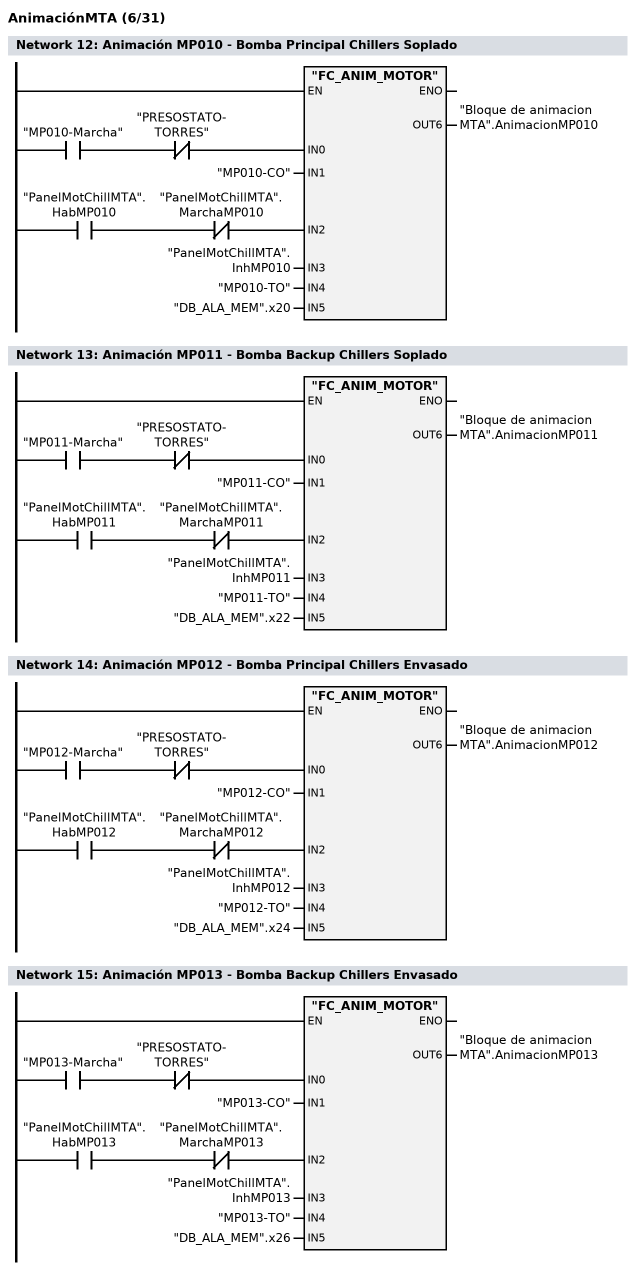
   RUNG wire#powerrail
      "FC_ANIM_MOTOR"(IN0 := wire#w1, IN2 := wire#w2, IN1 := "MP010-CO", IN3 := "PanelMotChillMTA".InhMP010, IN4 := "MP010-TO", IN5 := "DB_ALA_MEM".x20, OUT6 => "Bloque de animacion MTA".AnimacionMP010)
   END_RUNG
   RUNG wire#powerrail
      Contact( "MP010-Marcha" )
      I_Contact( "PRESOSTATO-TORRES" )
   END_RUNG wire#w1
   RUNG wire#powerrail
      Contact( "PanelMotChillMTA".HabMP010 )
      I_Contact( "PanelMotChillMTA".MarchaMP010 )
   END_RUNG wire#w2
   // the same network as SCL:
   "FC_ANIM_MOTOR"(IN0 := "MP010-Marcha" AND NOT "PRESOSTATO-TORRES",
                   IN1 := "MP010-CO",
                   IN2 := "PanelMotChillMTA".HabMP010 AND NOT "PanelMotChillMTA".MarchaMP010,
                   IN3 := "PanelMotChillMTA".InhMP010,
                   IN4 := "MP010-TO",
                   IN5 := "DB_ALA_MEM".x20,
                   OUT6 => "Bloque de animacion MTA".AnimacionMP010);
END_REGION

REGION Network 13: Animación MP011 - Bomba Backup Chillers Soplado
   RUNG wire#powerrail
      "FC_ANIM_MOTOR"(IN0 := wire#w1, IN2 := wire#w2, IN1 := "MP011-CO", IN3 := "PanelMotChillMTA".InhMP011, IN4 := "MP011-TO", IN5 := "DB_ALA_MEM".x22, OUT6 => "Bloque de animacion MTA".AnimacionMP011)
   END_RUNG
   RUNG wire#powerrail
      Contact( "MP011-Marcha" )
      I_Contact( "PRESOSTATO-TORRES" )
   END_RUNG wire#w1
   RUNG wire#powerrail
      Contact( "PanelMotChillMTA".HabMP011 )
      I_Contact( "PanelMotChillMTA".MarchaMP011 )
   END_RUNG wire#w2
   // the same network as SCL:
   "FC_ANIM_MOTOR"(IN0 := "MP011-Marcha" AND NOT "PRESOSTATO-TORRES",
                   IN1 := "MP011-CO",
                   IN2 := "PanelMotChillMTA".HabMP011 AND NOT "PanelMotChillMTA".MarchaMP011,
                   IN3 := "PanelMotChillMTA".InhMP011,
                   IN4 := "MP011-TO",
                   IN5 := "DB_ALA_MEM".x22,
                   OUT6 => "Bloque de animacion MTA".AnimacionMP011);
END_REGION

REGION Network 14: Animación MP012 - Bomba Principal Chillers Envasado
   RUNG wire#powerrail
      "FC_ANIM_MOTOR"(IN0 := wire#w1, IN2 := wire#w2, IN1 := "MP012-CO", IN3 := "PanelMotChillMTA".InhMP012, IN4 := "MP012-TO", IN5 := "DB_ALA_MEM".x24, OUT6 => "Bloque de animacion MTA".AnimacionMP012)
   END_RUNG
   RUNG wire#powerrail
      Contact( "MP012-Marcha" )
      I_Contact( "PRESOSTATO-TORRES" )
   END_RUNG wire#w1
   RUNG wire#powerrail
      Contact( "PanelMotChillMTA".HabMP012 )
      I_Contact( "PanelMotChillMTA".MarchaMP012 )
   END_RUNG wire#w2
   // the same network as SCL:
   "FC_ANIM_MOTOR"(IN0 := "MP012-Marcha" AND NOT "PRESOSTATO-TORRES",
                   IN1 := "MP012-CO",
                   IN2 := "PanelMotChillMTA".HabMP012 AND NOT "PanelMotChillMTA".MarchaMP012,
                   IN3 := "PanelMotChillMTA".InhMP012,
                   IN4 := "MP012-TO",
                   IN5 := "DB_ALA_MEM".x24,
                   OUT6 => "Bloque de animacion MTA".AnimacionMP012);
END_REGION

REGION Network 15: Animación MP013 - Bomba Backup Chillers Envasado
   RUNG wire#powerrail
      "FC_ANIM_MOTOR"(IN0 := wire#w1, IN2 := wire#w2, IN1 := "MP013-CO", IN3 := "PanelMotChillMTA".InhMP013, IN4 := "MP013-TO", IN5 := "DB_ALA_MEM".x26, OUT6 => "Bloque de animacion MTA".AnimacionMP013)
   END_RUNG
   RUNG wire#powerrail
      Contact( "MP013-Marcha" )
      I_Contact( "PRESOSTATO-TORRES" )
   END_RUNG wire#w1
   RUNG wire#powerrail
      Contact( "PanelMotChillMTA".HabMP013 )
      I_Contact( "PanelMotChillMTA".MarchaMP013 )
   END_RUNG wire#w2
   // the same network as SCL:
   "FC_ANIM_MOTOR"(IN0 := "MP013-Marcha" AND NOT "PRESOSTATO-TORRES",
                   IN1 := "MP013-CO",
                   IN2 := "PanelMotChillMTA".HabMP013 AND NOT "PanelMotChillMTA".MarchaMP013,
                   IN3 := "PanelMotChillMTA".InhMP013,
                   IN4 := "MP013-TO",
                   IN5 := "DB_ALA_MEM".x26,
                   OUT6 => "Bloque de animacion MTA".AnimacionMP013);
END_REGION

REGION Network 16: Animación MP018 - Bomba 1 Torres de enfriamiento
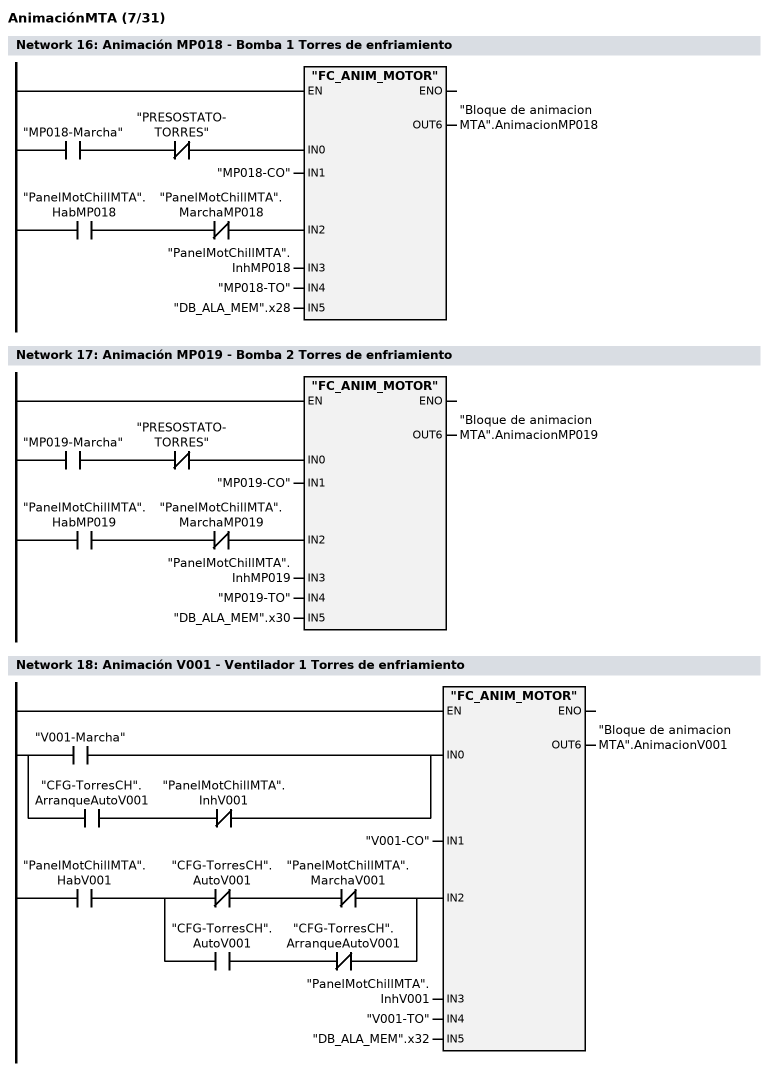
   RUNG wire#powerrail
      "FC_ANIM_MOTOR"(IN0 := wire#w1, IN2 := wire#w2, IN1 := "MP018-CO", IN3 := "PanelMotChillMTA".InhMP018, IN4 := "MP018-TO", IN5 := "DB_ALA_MEM".x28, OUT6 => "Bloque de animacion MTA".AnimacionMP018)
   END_RUNG
   RUNG wire#powerrail
      Contact( "MP018-Marcha" )
      I_Contact( "PRESOSTATO-TORRES" )
   END_RUNG wire#w1
   RUNG wire#powerrail
      Contact( "PanelMotChillMTA".HabMP018 )
      I_Contact( "PanelMotChillMTA".MarchaMP018 )
   END_RUNG wire#w2
   // the same network as SCL:
   "FC_ANIM_MOTOR"(IN0 := "MP018-Marcha" AND NOT "PRESOSTATO-TORRES",
                   IN1 := "MP018-CO",
                   IN2 := "PanelMotChillMTA".HabMP018 AND NOT "PanelMotChillMTA".MarchaMP018,
                   IN3 := "PanelMotChillMTA".InhMP018,
                   IN4 := "MP018-TO",
                   IN5 := "DB_ALA_MEM".x28,
                   OUT6 => "Bloque de animacion MTA".AnimacionMP018);
END_REGION

REGION Network 17: Animación MP019 - Bomba 2 Torres de enfriamiento
   RUNG wire#powerrail
      "FC_ANIM_MOTOR"(IN0 := wire#w1, IN2 := wire#w2, IN1 := "MP019-CO", IN3 := "PanelMotChillMTA".InhMP019, IN4 := "MP019-TO", IN5 := "DB_ALA_MEM".x30, OUT6 => "Bloque de animacion MTA".AnimacionMP019)
   END_RUNG
   RUNG wire#powerrail
      Contact( "MP019-Marcha" )
      I_Contact( "PRESOSTATO-TORRES" )
   END_RUNG wire#w1
   RUNG wire#powerrail
      Contact( "PanelMotChillMTA".HabMP019 )
      I_Contact( "PanelMotChillMTA".MarchaMP019 )
   END_RUNG wire#w2
   // the same network as SCL:
   "FC_ANIM_MOTOR"(IN0 := "MP019-Marcha" AND NOT "PRESOSTATO-TORRES",
                   IN1 := "MP019-CO",
                   IN2 := "PanelMotChillMTA".HabMP019 AND NOT "PanelMotChillMTA".MarchaMP019,
                   IN3 := "PanelMotChillMTA".InhMP019,
                   IN4 := "MP019-TO",
                   IN5 := "DB_ALA_MEM".x30,
                   OUT6 => "Bloque de animacion MTA".AnimacionMP019);
END_REGION

REGION Network 18: Animación V001 - Ventilador 1 Torres de enfriamiento
   RUNG wire#powerrail
      "FC_ANIM_MOTOR"(IN0 := wire#w1, IN2 := wire#w3, IN1 := "V001-CO", IN3 := "PanelMotChillMTA".InhV001, IN4 := "V001-TO", IN5 := "DB_ALA_MEM".x32, OUT6 => "Bloque de animacion MTA".AnimacionV001)
   END_RUNG
   RUNG wire#powerrail
      Contact( "V001-Marcha" )
   END_RUNG wire#w1
   RUNG wire#powerrail
      Contact( "CFG-TorresCH".ArranqueAutoV001 )
      I_Contact( "PanelMotChillMTA".InhV001 )
   END_RUNG wire#w1
   RUNG wire#powerrail
      Contact( "PanelMotChillMTA".HabV001 )
      wire#w2
      I_Contact( "CFG-TorresCH".AutoV001 )
      I_Contact( "PanelMotChillMTA".MarchaV001 )
   END_RUNG wire#w3
   RUNG wire#w2
      Contact( "CFG-TorresCH".AutoV001 )
      I_Contact( "CFG-TorresCH".ArranqueAutoV001 )
   END_RUNG wire#w3
   // the same network as SCL:
   "FC_ANIM_MOTOR"(IN0 := "V001-Marcha" OR ("CFG-TorresCH".ArranqueAutoV001 AND NOT "PanelMotChillMTA".InhV001),
                   IN1 := "V001-CO",
                   IN2 := "PanelMotChillMTA".HabV001 AND ((NOT "CFG-TorresCH".AutoV001 AND NOT "PanelMotChillMTA".MarchaV001) OR ("CFG-TorresCH".AutoV001 AND NOT "CFG-TorresCH".ArranqueAutoV001)),
                   IN3 := "PanelMotChillMTA".InhV001,
                   IN4 := "V001-TO",
                   IN5 := "DB_ALA_MEM".x32,
                   OUT6 => "Bloque de animacion MTA".AnimacionV001);
END_REGION

REGION Network 19: Animación V002 - Ventilador 2 Torres de enfriamiento
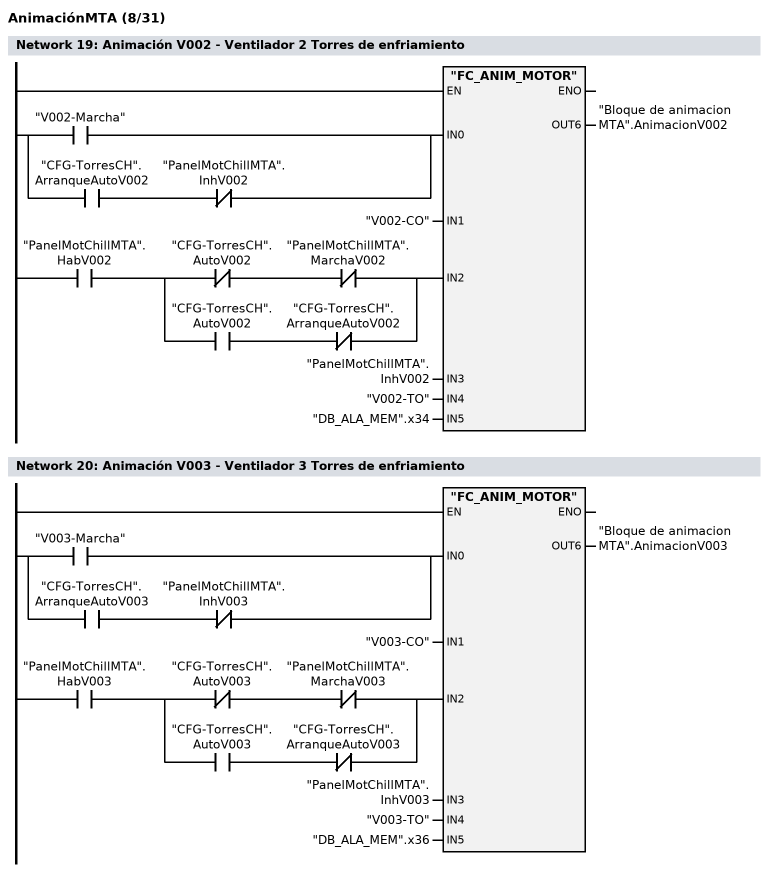
   RUNG wire#powerrail
      "FC_ANIM_MOTOR"(IN0 := wire#w1, IN2 := wire#w3, IN1 := "V002-CO", IN3 := "PanelMotChillMTA".InhV002, IN4 := "V002-TO", IN5 := "DB_ALA_MEM".x34, OUT6 => "Bloque de animacion MTA".AnimacionV002)
   END_RUNG
   RUNG wire#powerrail
      Contact( "V002-Marcha" )
   END_RUNG wire#w1
   RUNG wire#powerrail
      Contact( "CFG-TorresCH".ArranqueAutoV002 )
      I_Contact( "PanelMotChillMTA".InhV002 )
   END_RUNG wire#w1
   RUNG wire#powerrail
      Contact( "PanelMotChillMTA".HabV002 )
      wire#w2
      I_Contact( "CFG-TorresCH".AutoV002 )
      I_Contact( "PanelMotChillMTA".MarchaV002 )
   END_RUNG wire#w3
   RUNG wire#w2
      Contact( "CFG-TorresCH".AutoV002 )
      I_Contact( "CFG-TorresCH".ArranqueAutoV002 )
   END_RUNG wire#w3
   // the same network as SCL:
   "FC_ANIM_MOTOR"(IN0 := "V002-Marcha" OR ("CFG-TorresCH".ArranqueAutoV002 AND NOT "PanelMotChillMTA".InhV002),
                   IN1 := "V002-CO",
                   IN2 := "PanelMotChillMTA".HabV002 AND ((NOT "CFG-TorresCH".AutoV002 AND NOT "PanelMotChillMTA".MarchaV002) OR ("CFG-TorresCH".AutoV002 AND NOT "CFG-TorresCH".ArranqueAutoV002)),
                   IN3 := "PanelMotChillMTA".InhV002,
                   IN4 := "V002-TO",
                   IN5 := "DB_ALA_MEM".x34,
                   OUT6 => "Bloque de animacion MTA".AnimacionV002);
END_REGION

REGION Network 20: Animación V003 - Ventilador 3 Torres de enfriamiento
   RUNG wire#powerrail
      "FC_ANIM_MOTOR"(IN0 := wire#w1, IN2 := wire#w3, IN1 := "V003-CO", IN3 := "PanelMotChillMTA".InhV003, IN4 := "V003-TO", IN5 := "DB_ALA_MEM".x36, OUT6 => "Bloque de animacion MTA".AnimacionV003)
   END_RUNG
   RUNG wire#powerrail
      Contact( "V003-Marcha" )
   END_RUNG wire#w1
   RUNG wire#powerrail
      Contact( "CFG-TorresCH".ArranqueAutoV003 )
      I_Contact( "PanelMotChillMTA".InhV003 )
   END_RUNG wire#w1
   RUNG wire#powerrail
      Contact( "PanelMotChillMTA".HabV003 )
      wire#w2
      I_Contact( "CFG-TorresCH".AutoV003 )
      I_Contact( "PanelMotChillMTA".MarchaV003 )
   END_RUNG wire#w3
   RUNG wire#w2
      Contact( "CFG-TorresCH".AutoV003 )
      I_Contact( "CFG-TorresCH".ArranqueAutoV003 )
   END_RUNG wire#w3
   // the same network as SCL:
   "FC_ANIM_MOTOR"(IN0 := "V003-Marcha" OR ("CFG-TorresCH".ArranqueAutoV003 AND NOT "PanelMotChillMTA".InhV003),
                   IN1 := "V003-CO",
                   IN2 := "PanelMotChillMTA".HabV003 AND ((NOT "CFG-TorresCH".AutoV003 AND NOT "PanelMotChillMTA".MarchaV003) OR ("CFG-TorresCH".AutoV003 AND NOT "CFG-TorresCH".ArranqueAutoV003)),
                   IN3 := "PanelMotChillMTA".InhV003,
                   IN4 := "V003-TO",
                   IN5 := "DB_ALA_MEM".x36,
                   OUT6 => "Bloque de animacion MTA".AnimacionV003);
END_REGION

REGION Network 21: Animación MC060 - Compresor de Baja SULLAIR 2
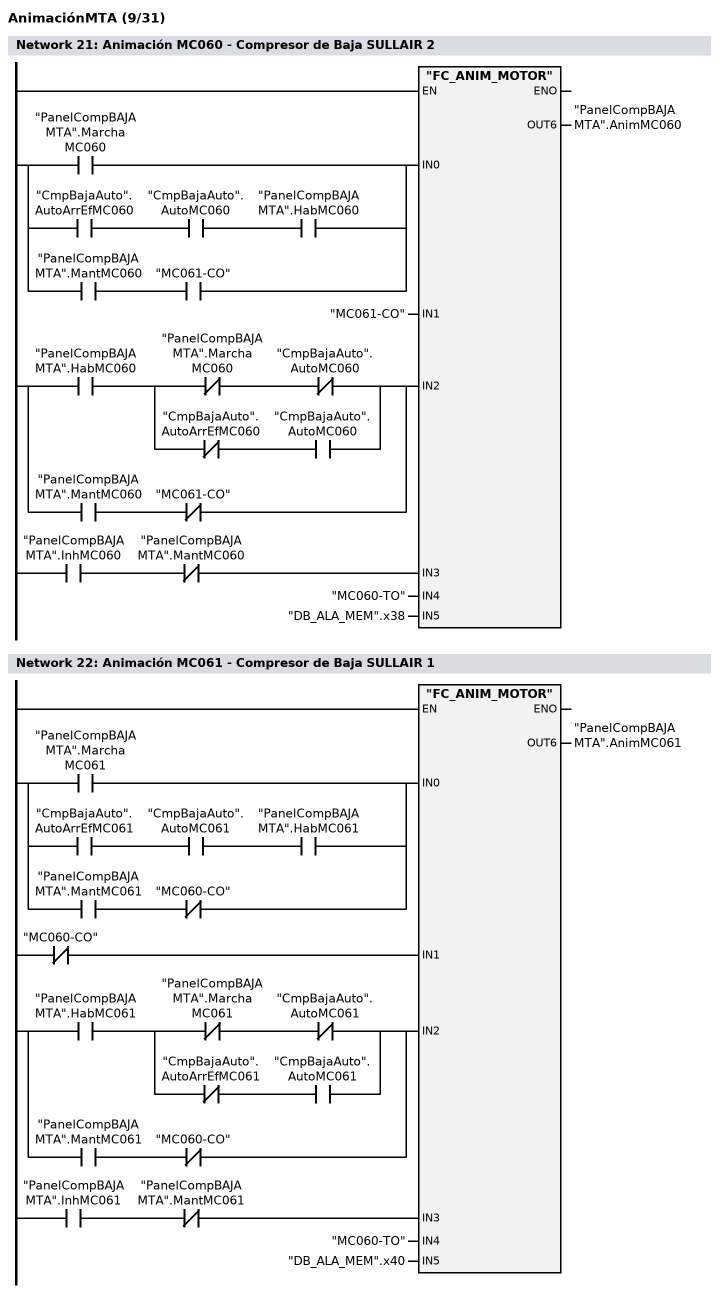
   RUNG wire#powerrail
      "FC_ANIM_MOTOR"(IN0 := wire#w1, IN2 := wire#w3, IN3 := wire#w4, IN1 := "MC061-CO", IN4 := "MC060-TO", IN5 := "DB_ALA_MEM".x38, OUT6 => "PanelCompBAJA MTA".AnimMC060)
   END_RUNG
   RUNG wire#powerrail
      Contact( "PanelCompBAJA MTA".MarchaMC060 )
   END_RUNG wire#w1
   RUNG wire#powerrail
      Contact( "CmpBajaAuto".AutoArrEfMC060 )
      Contact( "CmpBajaAuto".AutoMC060 )
      Contact( "PanelCompBAJA MTA".HabMC060 )
   END_RUNG wire#w1
   RUNG wire#powerrail
      Contact( "PanelCompBAJA MTA".MantMC060 )
      Contact( "MC061-CO" )
   END_RUNG wire#w1
   RUNG wire#powerrail
      Contact( "PanelCompBAJA MTA".HabMC060 )
      wire#w2
      I_Contact( "PanelCompBAJA MTA".MarchaMC060 )
      I_Contact( "CmpBajaAuto".AutoMC060 )
   END_RUNG wire#w3
   RUNG wire#w2
      I_Contact( "CmpBajaAuto".AutoArrEfMC060 )
      Contact( "CmpBajaAuto".AutoMC060 )
   END_RUNG wire#w3
   RUNG wire#powerrail
      Contact( "PanelCompBAJA MTA".MantMC060 )
      I_Contact( "MC061-CO" )
   END_RUNG wire#w3
   RUNG wire#powerrail
      Contact( "PanelCompBAJA MTA".InhMC060 )
      I_Contact( "PanelCompBAJA MTA".MantMC060 )
   END_RUNG wire#w4
   // the same network as SCL:
   "FC_ANIM_MOTOR"(IN0 := "PanelCompBAJA MTA".MarchaMC060 OR ("CmpBajaAuto".AutoArrEfMC060 AND "CmpBajaAuto".AutoMC060 AND "PanelCompBAJA MTA".HabMC060) OR ("PanelCompBAJA MTA".MantMC060 AND "MC061-CO"),
                   IN1 := "MC061-CO",
                   IN2 := ("PanelCompBAJA MTA".HabMC060 AND ((NOT "PanelCompBAJA MTA".MarchaMC060 AND NOT "CmpBajaAuto".AutoMC060) OR (NOT "CmpBajaAuto".AutoArrEfMC060 AND "CmpBajaAuto".AutoMC060))) OR ("PanelCompBAJA MTA".MantMC060 AND NOT "MC061-CO"),
                   IN3 := "PanelCompBAJA MTA".InhMC060 AND NOT "PanelCompBAJA MTA".MantMC060,
                   IN4 := "MC060-TO",
                   IN5 := "DB_ALA_MEM".x38,
                   OUT6 => "PanelCompBAJA MTA".AnimMC060);
END_REGION

REGION Network 22: Animación MC061 - Compresor de Baja SULLAIR 1
   RUNG wire#powerrail
      "FC_ANIM_MOTOR"(IN0 := wire#w1, IN1 := wire#w2, IN2 := wire#w4, IN3 := wire#w5, IN4 := "MC060-TO", IN5 := "DB_ALA_MEM".x40, OUT6 => "PanelCompBAJA MTA".AnimMC061)
   END_RUNG
   RUNG wire#powerrail
      Contact( "PanelCompBAJA MTA".MarchaMC061 )
   END_RUNG wire#w1
   RUNG wire#powerrail
      Contact( "CmpBajaAuto".AutoArrEfMC061 )
      Contact( "CmpBajaAuto".AutoMC061 )
      Contact( "PanelCompBAJA MTA".HabMC061 )
   END_RUNG wire#w1
   RUNG wire#powerrail
      Contact( "PanelCompBAJA MTA".MantMC061 )
      I_Contact( "MC060-CO" )
   END_RUNG wire#w1
   RUNG wire#powerrail
      I_Contact( "MC060-CO" )
   END_RUNG wire#w2
   RUNG wire#powerrail
      Contact( "PanelCompBAJA MTA".HabMC061 )
      wire#w3
      I_Contact( "PanelCompBAJA MTA".MarchaMC061 )
      I_Contact( "CmpBajaAuto".AutoMC061 )
   END_RUNG wire#w4
   RUNG wire#w3
      I_Contact( "CmpBajaAuto".AutoArrEfMC061 )
      Contact( "CmpBajaAuto".AutoMC061 )
   END_RUNG wire#w4
   RUNG wire#powerrail
      Contact( "PanelCompBAJA MTA".MantMC061 )
      I_Contact( "MC060-CO" )
   END_RUNG wire#w4
   RUNG wire#powerrail
      Contact( "PanelCompBAJA MTA".InhMC061 )
      I_Contact( "PanelCompBAJA MTA".MantMC061 )
   END_RUNG wire#w5
   // the same network as SCL:
   "FC_ANIM_MOTOR"(IN0 := "PanelCompBAJA MTA".MarchaMC061 OR ("CmpBajaAuto".AutoArrEfMC061 AND "CmpBajaAuto".AutoMC061 AND "PanelCompBAJA MTA".HabMC061) OR ("PanelCompBAJA MTA".MantMC061 AND NOT "MC060-CO"),
                   IN1 := NOT "MC060-CO",
                   IN2 := ("PanelCompBAJA MTA".HabMC061 AND ((NOT "PanelCompBAJA MTA".MarchaMC061 AND NOT "CmpBajaAuto".AutoMC061) OR (NOT "CmpBajaAuto".AutoArrEfMC061 AND "CmpBajaAuto".AutoMC061))) OR ("PanelCompBAJA MTA".MantMC061 AND NOT "MC060-CO"),
                   IN3 := "PanelCompBAJA MTA".InhMC061 AND NOT "PanelCompBAJA MTA".MantMC061,
                   IN4 := "MC060-TO",
                   IN5 := "DB_ALA_MEM".x40,
                   OUT6 => "PanelCompBAJA MTA".AnimMC061);
END_REGION

REGION Network 23: Animación MC062 - Compresor de Baja SULLAIR 0
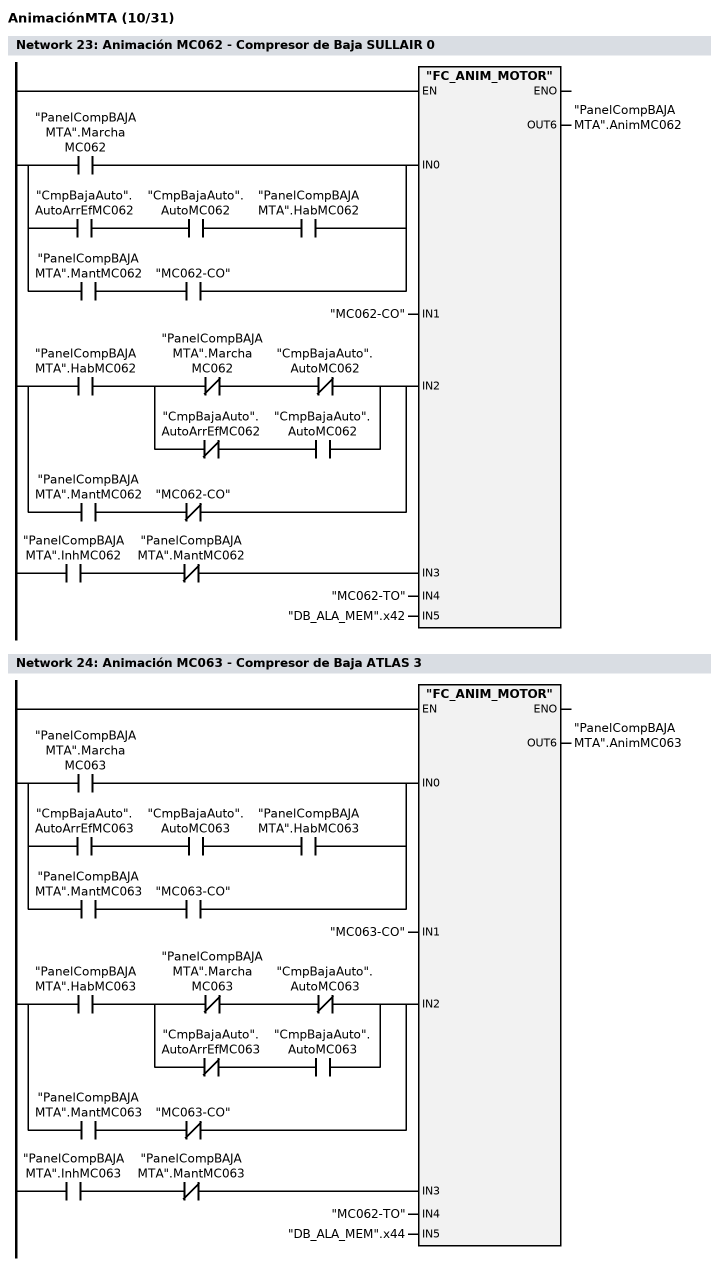
   RUNG wire#powerrail
      "FC_ANIM_MOTOR"(IN0 := wire#w1, IN2 := wire#w3, IN3 := wire#w4, IN1 := "MC062-CO", IN4 := "MC062-TO", IN5 := "DB_ALA_MEM".x42, OUT6 => "PanelCompBAJA MTA".AnimMC062)
   END_RUNG
   RUNG wire#powerrail
      Contact( "PanelCompBAJA MTA".MarchaMC062 )
   END_RUNG wire#w1
   RUNG wire#powerrail
      Contact( "CmpBajaAuto".AutoArrEfMC062 )
      Contact( "CmpBajaAuto".AutoMC062 )
      Contact( "PanelCompBAJA MTA".HabMC062 )
   END_RUNG wire#w1
   RUNG wire#powerrail
      Contact( "PanelCompBAJA MTA".MantMC062 )
      Contact( "MC062-CO" )
   END_RUNG wire#w1
   RUNG wire#powerrail
      Contact( "PanelCompBAJA MTA".HabMC062 )
      wire#w2
      I_Contact( "PanelCompBAJA MTA".MarchaMC062 )
      I_Contact( "CmpBajaAuto".AutoMC062 )
   END_RUNG wire#w3
   RUNG wire#w2
      I_Contact( "CmpBajaAuto".AutoArrEfMC062 )
      Contact( "CmpBajaAuto".AutoMC062 )
   END_RUNG wire#w3
   RUNG wire#powerrail
      Contact( "PanelCompBAJA MTA".MantMC062 )
      I_Contact( "MC062-CO" )
   END_RUNG wire#w3
   RUNG wire#powerrail
      Contact( "PanelCompBAJA MTA".InhMC062 )
      I_Contact( "PanelCompBAJA MTA".MantMC062 )
   END_RUNG wire#w4
   // the same network as SCL:
   "FC_ANIM_MOTOR"(IN0 := "PanelCompBAJA MTA".MarchaMC062 OR ("CmpBajaAuto".AutoArrEfMC062 AND "CmpBajaAuto".AutoMC062 AND "PanelCompBAJA MTA".HabMC062) OR ("PanelCompBAJA MTA".MantMC062 AND "MC062-CO"),
                   IN1 := "MC062-CO",
                   IN2 := ("PanelCompBAJA MTA".HabMC062 AND ((NOT "PanelCompBAJA MTA".MarchaMC062 AND NOT "CmpBajaAuto".AutoMC062) OR (NOT "CmpBajaAuto".AutoArrEfMC062 AND "CmpBajaAuto".AutoMC062))) OR ("PanelCompBAJA MTA".MantMC062 AND NOT "MC062-CO"),
                   IN3 := "PanelCompBAJA MTA".InhMC062 AND NOT "PanelCompBAJA MTA".MantMC062,
                   IN4 := "MC062-TO",
                   IN5 := "DB_ALA_MEM".x42,
                   OUT6 => "PanelCompBAJA MTA".AnimMC062);
END_REGION

REGION Network 24: Animación MC063 - Compresor de Baja ATLAS 3
   RUNG wire#powerrail
      "FC_ANIM_MOTOR"(IN0 := wire#w1, IN2 := wire#w3, IN3 := wire#w4, IN1 := "MC063-CO", IN4 := "MC062-TO", IN5 := "DB_ALA_MEM".x44, OUT6 => "PanelCompBAJA MTA".AnimMC063)
   END_RUNG
   RUNG wire#powerrail
      Contact( "PanelCompBAJA MTA".MarchaMC063 )
   END_RUNG wire#w1
   RUNG wire#powerrail
      Contact( "CmpBajaAuto".AutoArrEfMC063 )
      Contact( "CmpBajaAuto".AutoMC063 )
      Contact( "PanelCompBAJA MTA".HabMC063 )
   END_RUNG wire#w1
   RUNG wire#powerrail
      Contact( "PanelCompBAJA MTA".MantMC063 )
      Contact( "MC063-CO" )
   END_RUNG wire#w1
   RUNG wire#powerrail
      Contact( "PanelCompBAJA MTA".HabMC063 )
      wire#w2
      I_Contact( "PanelCompBAJA MTA".MarchaMC063 )
      I_Contact( "CmpBajaAuto".AutoMC063 )
   END_RUNG wire#w3
   RUNG wire#w2
      I_Contact( "CmpBajaAuto".AutoArrEfMC063 )
      Contact( "CmpBajaAuto".AutoMC063 )
   END_RUNG wire#w3
   RUNG wire#powerrail
      Contact( "PanelCompBAJA MTA".MantMC063 )
      I_Contact( "MC063-CO" )
   END_RUNG wire#w3
   RUNG wire#powerrail
      Contact( "PanelCompBAJA MTA".InhMC063 )
      I_Contact( "PanelCompBAJA MTA".MantMC063 )
   END_RUNG wire#w4
   // the same network as SCL:
   "FC_ANIM_MOTOR"(IN0 := "PanelCompBAJA MTA".MarchaMC063 OR ("CmpBajaAuto".AutoArrEfMC063 AND "CmpBajaAuto".AutoMC063 AND "PanelCompBAJA MTA".HabMC063) OR ("PanelCompBAJA MTA".MantMC063 AND "MC063-CO"),
                   IN1 := "MC063-CO",
                   IN2 := ("PanelCompBAJA MTA".HabMC063 AND ((NOT "PanelCompBAJA MTA".MarchaMC063 AND NOT "CmpBajaAuto".AutoMC063) OR (NOT "CmpBajaAuto".AutoArrEfMC063 AND "CmpBajaAuto".AutoMC063))) OR ("PanelCompBAJA MTA".MantMC063 AND NOT "MC063-CO"),
                   IN3 := "PanelCompBAJA MTA".InhMC063 AND NOT "PanelCompBAJA MTA".MantMC063,
                   IN4 := "MC062-TO",
                   IN5 := "DB_ALA_MEM".x44,
                   OUT6 => "PanelCompBAJA MTA".AnimMC063);
END_REGION

REGION Network 25: Animación MC064 - Compresor de Baja ATLAS 2
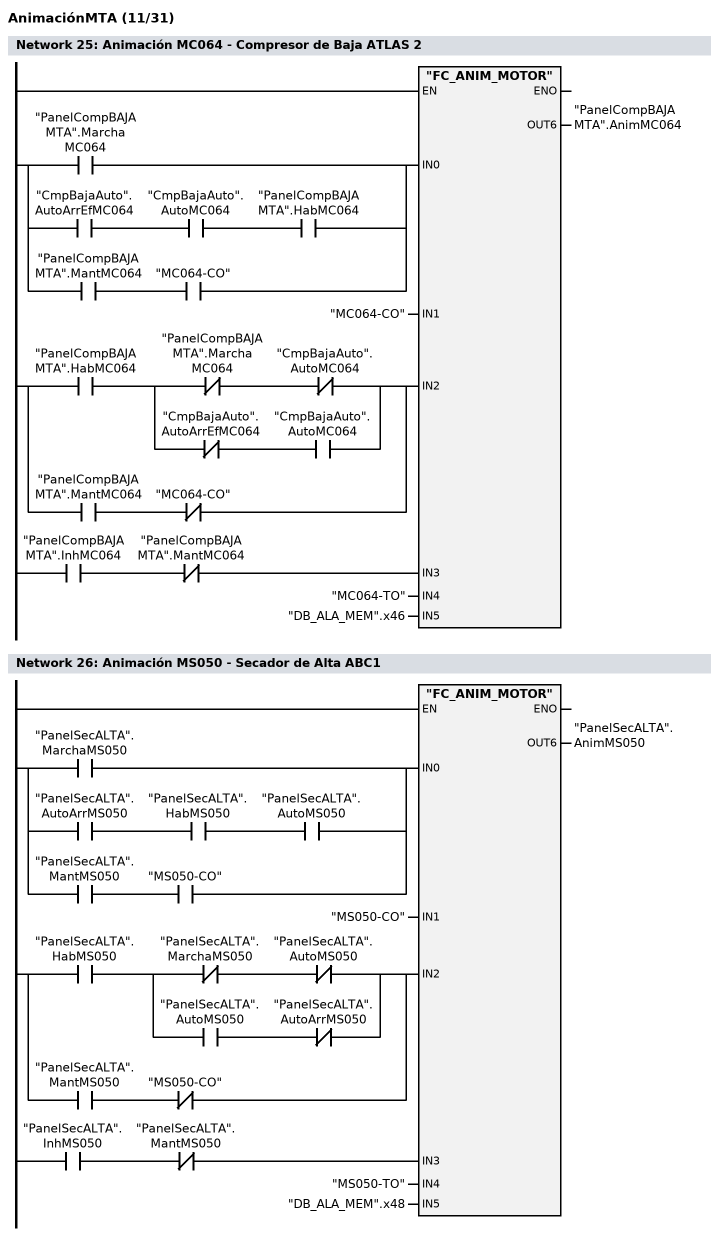
   RUNG wire#powerrail
      "FC_ANIM_MOTOR"(IN0 := wire#w1, IN2 := wire#w3, IN3 := wire#w4, IN1 := "MC064-CO", IN4 := "MC064-TO", IN5 := "DB_ALA_MEM".x46, OUT6 => "PanelCompBAJA MTA".AnimMC064)
   END_RUNG
   RUNG wire#powerrail
      Contact( "PanelCompBAJA MTA".MarchaMC064 )
   END_RUNG wire#w1
   RUNG wire#powerrail
      Contact( "CmpBajaAuto".AutoArrEfMC064 )
      Contact( "CmpBajaAuto".AutoMC064 )
      Contact( "PanelCompBAJA MTA".HabMC064 )
   END_RUNG wire#w1
   RUNG wire#powerrail
      Contact( "PanelCompBAJA MTA".MantMC064 )
      Contact( "MC064-CO" )
   END_RUNG wire#w1
   RUNG wire#powerrail
      Contact( "PanelCompBAJA MTA".HabMC064 )
      wire#w2
      I_Contact( "PanelCompBAJA MTA".MarchaMC064 )
      I_Contact( "CmpBajaAuto".AutoMC064 )
   END_RUNG wire#w3
   RUNG wire#w2
      I_Contact( "CmpBajaAuto".AutoArrEfMC064 )
      Contact( "CmpBajaAuto".AutoMC064 )
   END_RUNG wire#w3
   RUNG wire#powerrail
      Contact( "PanelCompBAJA MTA".MantMC064 )
      I_Contact( "MC064-CO" )
   END_RUNG wire#w3
   RUNG wire#powerrail
      Contact( "PanelCompBAJA MTA".InhMC064 )
      I_Contact( "PanelCompBAJA MTA".MantMC064 )
   END_RUNG wire#w4
   // the same network as SCL:
   "FC_ANIM_MOTOR"(IN0 := "PanelCompBAJA MTA".MarchaMC064 OR ("CmpBajaAuto".AutoArrEfMC064 AND "CmpBajaAuto".AutoMC064 AND "PanelCompBAJA MTA".HabMC064) OR ("PanelCompBAJA MTA".MantMC064 AND "MC064-CO"),
                   IN1 := "MC064-CO",
                   IN2 := ("PanelCompBAJA MTA".HabMC064 AND ((NOT "PanelCompBAJA MTA".MarchaMC064 AND NOT "CmpBajaAuto".AutoMC064) OR (NOT "CmpBajaAuto".AutoArrEfMC064 AND "CmpBajaAuto".AutoMC064))) OR ("PanelCompBAJA MTA".MantMC064 AND NOT "MC064-CO"),
                   IN3 := "PanelCompBAJA MTA".InhMC064 AND NOT "PanelCompBAJA MTA".MantMC064,
                   IN4 := "MC064-TO",
                   IN5 := "DB_ALA_MEM".x46,
                   OUT6 => "PanelCompBAJA MTA".AnimMC064);
END_REGION

REGION Network 26: Animación MS050 - Secador de Alta ABC1
   RUNG wire#powerrail
      "FC_ANIM_MOTOR"(IN0 := wire#w1, IN2 := wire#w3, IN3 := wire#w4, IN1 := "MS050-CO", IN4 := "MS050-TO", IN5 := "DB_ALA_MEM".x48, OUT6 => "PanelSecALTA".AnimMS050)
   END_RUNG
   RUNG wire#powerrail
      Contact( "PanelSecALTA".MarchaMS050 )
   END_RUNG wire#w1
   RUNG wire#powerrail
      Contact( "PanelSecALTA".AutoArrMS050 )
      Contact( "PanelSecALTA".HabMS050 )
      Contact( "PanelSecALTA".AutoMS050 )
   END_RUNG wire#w1
   RUNG wire#powerrail
      Contact( "PanelSecALTA".MantMS050 )
      Contact( "MS050-CO" )
   END_RUNG wire#w1
   RUNG wire#powerrail
      Contact( "PanelSecALTA".HabMS050 )
      wire#w2
      I_Contact( "PanelSecALTA".MarchaMS050 )
      I_Contact( "PanelSecALTA".AutoMS050 )
   END_RUNG wire#w3
   RUNG wire#w2
      Contact( "PanelSecALTA".AutoMS050 )
      I_Contact( "PanelSecALTA".AutoArrMS050 )
   END_RUNG wire#w3
   RUNG wire#powerrail
      Contact( "PanelSecALTA".MantMS050 )
      I_Contact( "MS050-CO" )
   END_RUNG wire#w3
   RUNG wire#powerrail
      Contact( "PanelSecALTA".InhMS050 )
      I_Contact( "PanelSecALTA".MantMS050 )
   END_RUNG wire#w4
   // the same network as SCL:
   "FC_ANIM_MOTOR"(IN0 := "PanelSecALTA".MarchaMS050 OR ("PanelSecALTA".AutoArrMS050 AND "PanelSecALTA".HabMS050 AND "PanelSecALTA".AutoMS050) OR ("PanelSecALTA".MantMS050 AND "MS050-CO"),
                   IN1 := "MS050-CO",
                   IN2 := ("PanelSecALTA".HabMS050 AND ((NOT "PanelSecALTA".MarchaMS050 AND NOT "PanelSecALTA".AutoMS050) OR ("PanelSecALTA".AutoMS050 AND NOT "PanelSecALTA".AutoArrMS050))) OR ("PanelSecALTA".MantMS050 AND NOT "MS050-CO"),
                   IN3 := "PanelSecALTA".InhMS050 AND NOT "PanelSecALTA".MantMS050,
                   IN4 := "MS050-TO",
                   IN5 := "DB_ALA_MEM".x48,
                   OUT6 => "PanelSecALTA".AnimMS050);
END_REGION

REGION Network 27: Animación MS051 - Secador de Alta ABC3
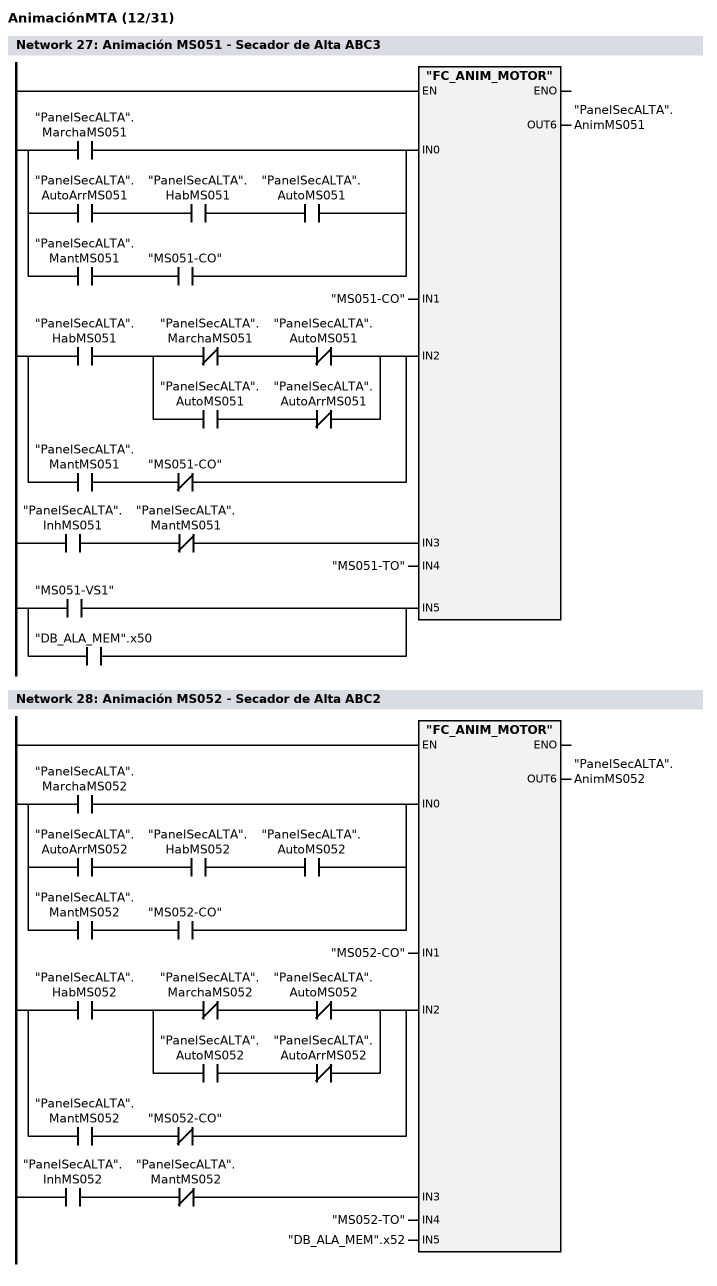
   RUNG wire#powerrail
      "FC_ANIM_MOTOR"(IN0 := wire#w1, IN2 := wire#w3, IN3 := wire#w4, IN5 := wire#w5, IN1 := "MS051-CO", IN4 := "MS051-TO", OUT6 => "PanelSecALTA".AnimMS051)
   END_RUNG
   RUNG wire#powerrail
      Contact( "PanelSecALTA".MarchaMS051 )
   END_RUNG wire#w1
   RUNG wire#powerrail
      Contact( "PanelSecALTA".AutoArrMS051 )
      Contact( "PanelSecALTA".HabMS051 )
      Contact( "PanelSecALTA".AutoMS051 )
   END_RUNG wire#w1
   RUNG wire#powerrail
      Contact( "PanelSecALTA".MantMS051 )
      Contact( "MS051-CO" )
   END_RUNG wire#w1
   RUNG wire#powerrail
      Contact( "PanelSecALTA".HabMS051 )
      wire#w2
      I_Contact( "PanelSecALTA".MarchaMS051 )
      I_Contact( "PanelSecALTA".AutoMS051 )
   END_RUNG wire#w3
   RUNG wire#w2
      Contact( "PanelSecALTA".AutoMS051 )
      I_Contact( "PanelSecALTA".AutoArrMS051 )
   END_RUNG wire#w3
   RUNG wire#powerrail
      Contact( "PanelSecALTA".MantMS051 )
      I_Contact( "MS051-CO" )
   END_RUNG wire#w3
   RUNG wire#powerrail
      Contact( "PanelSecALTA".InhMS051 )
      I_Contact( "PanelSecALTA".MantMS051 )
   END_RUNG wire#w4
   RUNG wire#powerrail
      Contact( "MS051-VS1" )
   END_RUNG wire#w5
   RUNG wire#powerrail
      Contact( "DB_ALA_MEM".x50 )
   END_RUNG wire#w5
   // the same network as SCL:
   "FC_ANIM_MOTOR"(IN0 := "PanelSecALTA".MarchaMS051 OR ("PanelSecALTA".AutoArrMS051 AND "PanelSecALTA".HabMS051 AND "PanelSecALTA".AutoMS051) OR ("PanelSecALTA".MantMS051 AND "MS051-CO"),
                   IN1 := "MS051-CO",
                   IN2 := ("PanelSecALTA".HabMS051 AND ((NOT "PanelSecALTA".MarchaMS051 AND NOT "PanelSecALTA".AutoMS051) OR ("PanelSecALTA".AutoMS051 AND NOT "PanelSecALTA".AutoArrMS051))) OR ("PanelSecALTA".MantMS051 AND NOT "MS051-CO"),
                   IN3 := "PanelSecALTA".InhMS051 AND NOT "PanelSecALTA".MantMS051,
                   IN4 := "MS051-TO",
                   IN5 := "MS051-VS1" OR "DB_ALA_MEM".x50,
                   OUT6 => "PanelSecALTA".AnimMS051);
END_REGION

REGION Network 28: Animación MS052 - Secador de Alta ABC2
   RUNG wire#powerrail
      "FC_ANIM_MOTOR"(IN0 := wire#w1, IN2 := wire#w3, IN3 := wire#w4, IN1 := "MS052-CO", IN4 := "MS052-TO", IN5 := "DB_ALA_MEM".x52, OUT6 => "PanelSecALTA".AnimMS052)
   END_RUNG
   RUNG wire#powerrail
      Contact( "PanelSecALTA".MarchaMS052 )
   END_RUNG wire#w1
   RUNG wire#powerrail
      Contact( "PanelSecALTA".AutoArrMS052 )
      Contact( "PanelSecALTA".HabMS052 )
      Contact( "PanelSecALTA".AutoMS052 )
   END_RUNG wire#w1
   RUNG wire#powerrail
      Contact( "PanelSecALTA".MantMS052 )
      Contact( "MS052-CO" )
   END_RUNG wire#w1
   RUNG wire#powerrail
      Contact( "PanelSecALTA".HabMS052 )
      wire#w2
      I_Contact( "PanelSecALTA".MarchaMS052 )
      I_Contact( "PanelSecALTA".AutoMS052 )
   END_RUNG wire#w3
   RUNG wire#w2
      Contact( "PanelSecALTA".AutoMS052 )
      I_Contact( "PanelSecALTA".AutoArrMS052 )
   END_RUNG wire#w3
   RUNG wire#powerrail
      Contact( "PanelSecALTA".MantMS052 )
      I_Contact( "MS052-CO" )
   END_RUNG wire#w3
   RUNG wire#powerrail
      Contact( "PanelSecALTA".InhMS052 )
      I_Contact( "PanelSecALTA".MantMS052 )
   END_RUNG wire#w4
   // the same network as SCL:
   "FC_ANIM_MOTOR"(IN0 := "PanelSecALTA".MarchaMS052 OR ("PanelSecALTA".AutoArrMS052 AND "PanelSecALTA".HabMS052 AND "PanelSecALTA".AutoMS052) OR ("PanelSecALTA".MantMS052 AND "MS052-CO"),
                   IN1 := "MS052-CO",
                   IN2 := ("PanelSecALTA".HabMS052 AND ((NOT "PanelSecALTA".MarchaMS052 AND NOT "PanelSecALTA".AutoMS052) OR ("PanelSecALTA".AutoMS052 AND NOT "PanelSecALTA".AutoArrMS052))) OR ("PanelSecALTA".MantMS052 AND NOT "MS052-CO"),
                   IN3 := "PanelSecALTA".InhMS052 AND NOT "PanelSecALTA".MantMS052,
                   IN4 := "MS052-TO",
                   IN5 := "DB_ALA_MEM".x52,
                   OUT6 => "PanelSecALTA".AnimMS052);
END_REGION

REGION Network 29: Animación MS053 - Secador de Alta FARGON
